REGION Network 16: TBD Stacking_New : Control Balize
   RUNG wire#powerrail
      Contact( "DB_MDM_SN".Energie )
      wire#w1
      Coil( #SN_bsr )
      Coil( "SN_Baliza dulap rosu" )
   END_RUNG
   RUNG wire#powerrail
      Contact( "DB_MDM_SN".No_Safe )
   END_RUNG wire#w1
   RUNG wire#powerrail
      Contact( "Gen".SN_AlarmAny )
   END_RUNG wire#w1
   RUNG wire#powerrail
      { S7_Templates := "SrcType := USInt" } EQ_Contact(in1 := "sn".f[5]."step", in2 := 2)
      wire#w2
      Contact( "DB2_WORK_BITS".Stacker_New_Handler.Input.Vertical_sus )
      Contact( "DB2_WORK_BITS".Stacker_New_Handler.Input.Furca_extins )
      Coil( #SN_bsy )
   END_RUNG
   RUNG wire#powerrail
      { S7_Templates := "SrcType := USInt" } EQ_Contact(in1 := "sn".f[5]."step", in2 := 4)
   END_RUNG wire#w2
   RUNG wire#powerrail
      I_Contact( "DB_MDM_SN".Energie )
      I_Contact( "DB_MDM_SN".No_Safe )
      I_Contact( "DB_MDM_SN".Cycle_Run )
      Coil( #SN_bsgc )
   END_RUNG
   RUNG wire#powerrail
      Contact( #SN_bsgc )
      Contact( "Clock_0.5Hz" )
      wire#w3
      Coil( "Sn_Baliza dulap verde" )
   END_RUNG
   RUNG wire#powerrail
      Contact( "DB_MDM_SN".Cycle_Run )
   END_RUNG wire#w3
   RUNG wire#w3
      Coil( #SN_bsg )
   END_RUNG
   RUNG wire#powerrail
      Contact( #SN_bsg )
      I_Contact( #SN_bsgc )
      Contact( #SN_bsy )
      Contact( "Clock_0.5Hz" )
      wire#w4
      Coil( "BS_G" )
   END_RUNG
   RUNG wire#powerrail
      Contact( #SN_bsg )
      I_Contact( #SN_bsy )
   END_RUNG wire#w4
   RUNG wire#powerrail
      Contact( #SN_bsg )
      Contact( #SN_bsy )
      wire#w5
      I_Contact( "Clock_0.5Hz" )
      Coil( "BS_Y" )
   END_RUNG
   RUNG wire#powerrail
      Contact( #SN_bsgc )
      Contact( #SN_bsy )
   END_RUNG wire#w5
   RUNG wire#powerrail
      Contact( #SN_bsr )
      Contact( #SN_bsy )
   END_RUNG wire#w5
   RUNG wire#powerrail
      Contact( #SN_bsr )
      wire#w6
      Contact( #SN_bsy )
      Contact( "Clock_0.5Hz" )
      wire#w7
      Coil( "BS_R" )
   END_RUNG
   RUNG wire#w6
      I_Contact( #SN_bsy )
   END_RUNG wire#w7
   // the same network as SCL:
   #SN_bsr := "DB_MDM_SN".Energie OR "DB_MDM_SN".No_Safe OR "Gen".SN_AlarmAny;
   "SN_Baliza dulap rosu" := #SN_bsr;
   #SN_bsy := (("sn".f[5]."step" = 2) OR ("sn".f[5]."step" = 4)) AND "DB2_WORK_BITS".Stacker_New_Handler.Input.Vertical_sus AND "DB2_WORK_BITS".Stacker_New_Handler.Input.Furca_extins;
   #SN_bsgc := NOT "DB_MDM_SN".Energie AND NOT "DB_MDM_SN".No_Safe AND NOT "DB_MDM_SN".Cycle_Run;
   "Sn_Baliza dulap verde" := (#SN_bsgc AND "Clock_0.5Hz") OR "DB_MDM_SN".Cycle_Run;
   #SN_bsg := "Sn_Baliza dulap verde";
   "BS_G" := (#SN_bsg AND NOT #SN_bsgc AND #SN_bsy AND "Clock_0.5Hz") OR (#SN_bsg AND NOT #SN_bsy);
   "BS_Y" := ((#SN_bsg AND #SN_bsy) OR (#SN_bsgc AND #SN_bsy) OR (#SN_bsr AND #SN_bsy)) AND NOT "Clock_0.5Hz";
   "BS_R" := #SN_bsr AND ((#SN_bsy AND "Clock_0.5Hz") OR NOT #SN_bsy);
END_REGION
END_FUNCTION

FUNCTION "FC20_HMI" : Void   // FC20, LAD
{ S7_Optimized_Access := 'TRUE' }
VERSION : 0.1
BEGIN

REGION Network 1
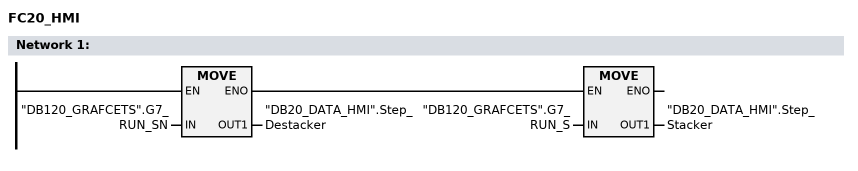
   RUNG wire#powerrail
      Move(in := "DB120_GRAFCETS".G7_RUN_SN, out1 => "DB20_DATA_HMI".Step_Destacker)
      Move(in := "DB120_GRAFCETS".G7_RUN_S, out1 => "DB20_DATA_HMI".Step_Stacker)
   END_RUNG
   // the same network as SCL:
   "DB20_DATA_HMI".Step_Destacker := "DB120_GRAFCETS".G7_RUN_SN;
   "DB20_DATA_HMI".Step_Stacker := "DB120_GRAFCETS".G7_RUN_S;
END_REGION
END_FUNCTION

FUNCTION "FC52_STACKING_New" : Void   // FC49, LAD
{ S7_Optimized_Access := 'TRUE' }
VERSION : 0.1
   VAR_TEMP
      Reset_S_Up : Bool;
      Reset_S_Fork : Bool;
      iB5_p : Bool;
      Reset_S : Bool;
      dumyb : Bool;
      dumyw : Int;
   END_VAR
   VAR_TEMP   // added for the SCL form of the ladder/FBD networks
      _w1 : Bool;
      _w2 : Bool;
      _w3 : Bool;
   END_VAR
BEGIN

REGION Network 1: mdm
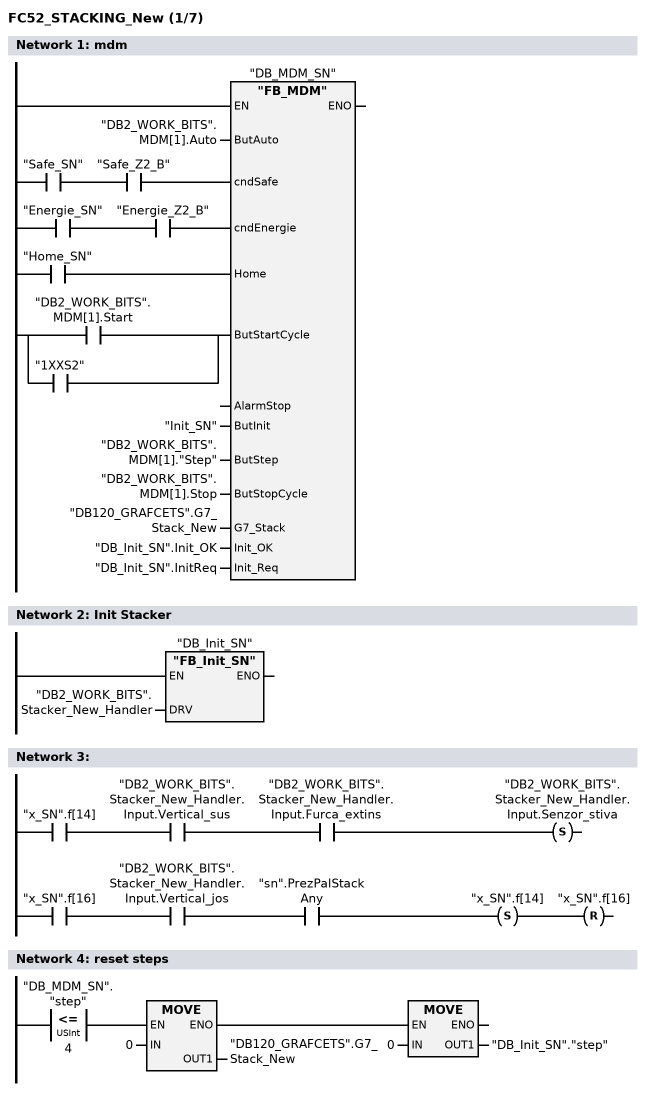
   RUNG wire#powerrail
      "DB_MDM_SN"(cndSafe := wire#w1, cndEnergie := wire#w2, Home := wire#w3, ButStartCycle := wire#w4, ButAuto := "DB2_WORK_BITS".MDM[1].Auto, AlarmStop :=, ButInit := "Init_SN", ButStep := "DB2_WORK_BITS".MDM[1]."Step", ButStopCycle := "DB2_WORK_BITS".MDM[1].Stop, G7_Stack := "DB120_GRAFCETS".G7_Stack_New, Init_OK := "DB_Init_SN".Init_OK, Init_Req := "DB_Init_SN".InitReq)
   END_RUNG
   RUNG wire#powerrail
      Contact( "Safe_SN" )
      Contact( "Safe_Z2_B" )
   END_RUNG wire#w1
   RUNG wire#powerrail
      Contact( "Energie_SN" )
      Contact( "Energie_Z2_B" )
   END_RUNG wire#w2
   RUNG wire#powerrail
      Contact( "Home_SN" )
   END_RUNG wire#w3
   RUNG wire#powerrail
      Contact( "DB2_WORK_BITS".MDM[1].Start )
   END_RUNG wire#w4
   RUNG wire#powerrail
      Contact( "1XXS2" )
   END_RUNG wire#w4
   // the same network as SCL:
   "DB_MDM_SN"(ButAuto := "DB2_WORK_BITS".MDM[1].Auto,   // "FB_MDM"
               cndSafe := "Safe_SN" AND "Safe_Z2_B",
               cndEnergie := "Energie_SN" AND "Energie_Z2_B",
               Home := "Home_SN",
               ButStartCycle := "DB2_WORK_BITS".MDM[1].Start OR "1XXS2",
               ButInit := "Init_SN",
               ButStep := "DB2_WORK_BITS".MDM[1]."Step",
               ButStopCycle := "DB2_WORK_BITS".MDM[1].Stop,
               G7_Stack := "DB120_GRAFCETS".G7_Stack_New,
               Init_OK := "DB_Init_SN".Init_OK,
               Init_Req := "DB_Init_SN".InitReq);
END_REGION

REGION Network 2: Init Stacker
   RUNG wire#powerrail
      "DB_Init_SN"(DRV := "DB2_WORK_BITS".Stacker_New_Handler)
   END_RUNG
   // the same network as SCL:
   "DB_Init_SN"(DRV := "DB2_WORK_BITS".Stacker_New_Handler);   // "FB_Init_SN"
END_REGION

REGION Network 3
   RUNG wire#powerrail
      Contact( "x_SN".f[14] )
      Contact( "DB2_WORK_BITS".Stacker_New_Handler.Input.Vertical_sus )
      Contact( "DB2_WORK_BITS".Stacker_New_Handler.Input.Furca_extins )
      S_Coil( "DB2_WORK_BITS".Stacker_New_Handler.Input.Senzor_stiva )
   END_RUNG
   RUNG wire#powerrail
      Contact( "x_SN".f[16] )
      Contact( "DB2_WORK_BITS".Stacker_New_Handler.Input.Vertical_jos )
      Contact( "sn".PrezPalStackAny )
      S_Coil( "x_SN".f[14] )
      R_Coil( "x_SN".f[16] )
   END_RUNG
   // the same network as SCL:
   IF "x_SN".f[14] AND "DB2_WORK_BITS".Stacker_New_Handler.Input.Vertical_sus AND "DB2_WORK_BITS".Stacker_New_Handler.Input.Furca_extins THEN
       "DB2_WORK_BITS".Stacker_New_Handler.Input.Senzor_stiva := TRUE;
   END_IF;
   #_w1 := "x_SN".f[16] AND "DB2_WORK_BITS".Stacker_New_Handler.Input.Vertical_jos AND "sn".PrezPalStackAny;
   IF #_w1 THEN
       "x_SN".f[14] := TRUE;
       "x_SN".f[16] := FALSE;
   END_IF;
END_REGION

REGION Network 4: reset steps
   RUNG wire#powerrail
      { S7_Templates := "SrcType := USInt" } LE_Contact(in1 := "DB_MDM_SN"."step", in2 := 4)
      Move(in := 0, out1 => "DB120_GRAFCETS".G7_Stack_New)
      Move(in := 0, out1 => "DB_Init_SN"."step")
   END_RUNG
   // the same network as SCL:
   IF "DB_MDM_SN"."step" <= 4 THEN
       "DB120_GRAFCETS".G7_Stack_New := 0;
       "DB_Init_SN"."step" := 0;
   END_IF;
END_REGION

REGION Network 5: start graf stack
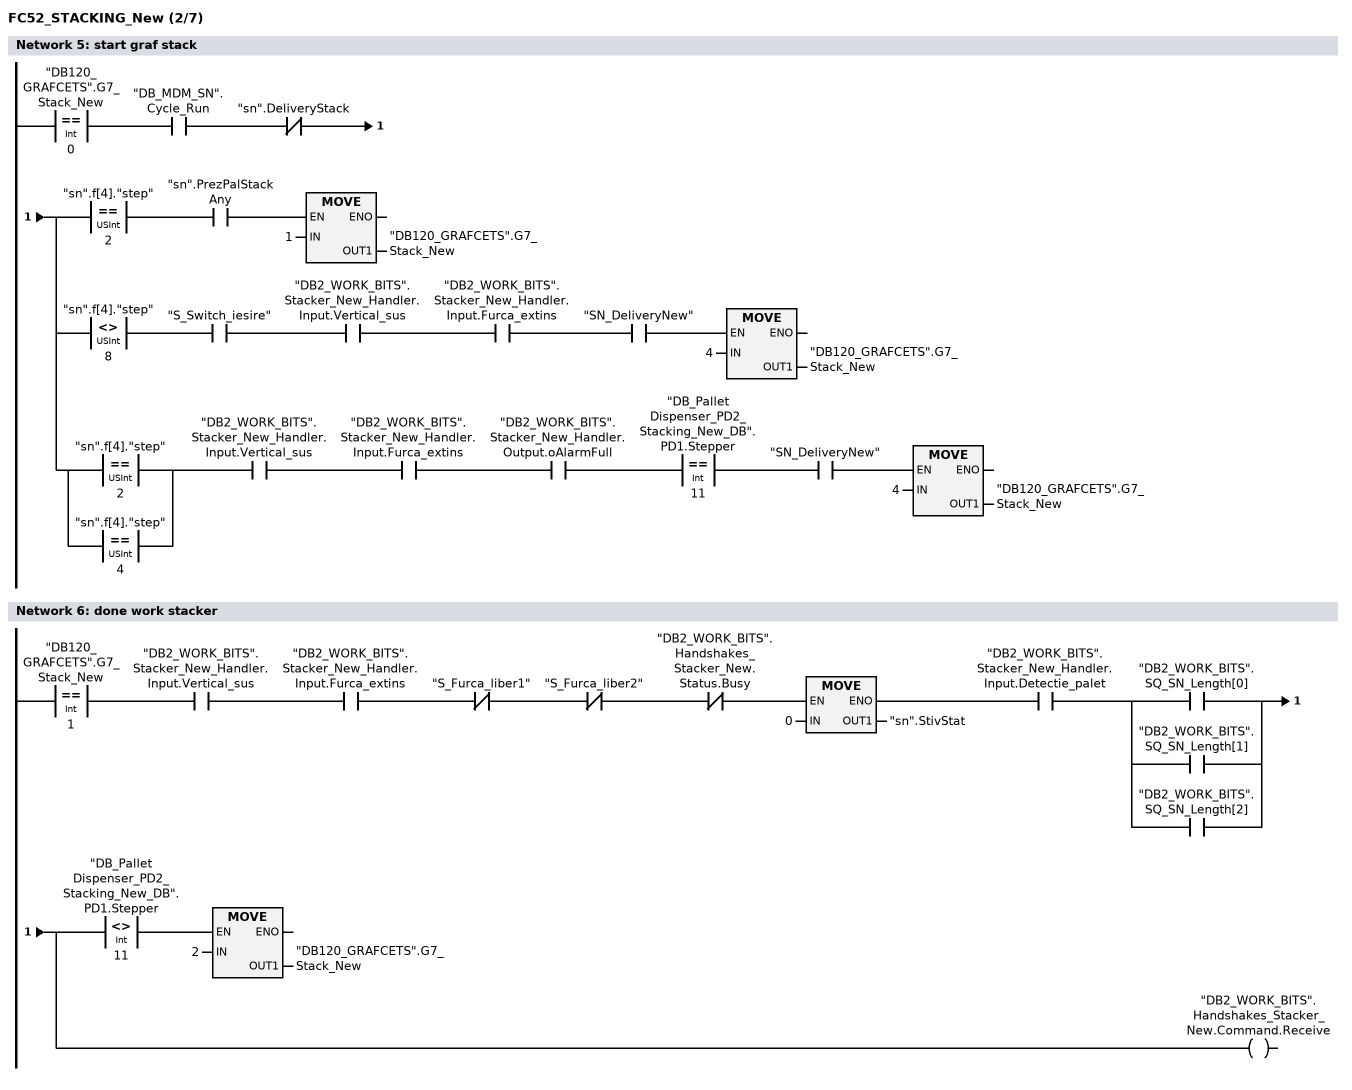
   RUNG wire#powerrail
      { S7_Templates := "SrcType := Int" } EQ_Contact(in1 := "DB120_GRAFCETS".G7_Stack_New, in2 := 0)
      Contact( "DB_MDM_SN".Cycle_Run )
      I_Contact( "sn".DeliveryStack )
      wire#w1
      { S7_Templates := "SrcType := USInt" } EQ_Contact(in1 := "sn".f[4]."step", in2 := 2)
      Contact( "sn".PrezPalStackAny )
      Move(in := 1, out1 => "DB120_GRAFCETS".G7_Stack_New)
   END_RUNG
   RUNG wire#w1
      { S7_Templates := "SrcType := USInt" } NE_Contact(in1 := "sn".f[4]."step", in2 := 8)
      Contact( "S_Switch_iesire" )
      Contact( "DB2_WORK_BITS".Stacker_New_Handler.Input.Vertical_sus )
      Contact( "DB2_WORK_BITS".Stacker_New_Handler.Input.Furca_extins )
      Contact( "SN_DeliveryNew" )
      Move(in := 4, out1 => "DB120_GRAFCETS".G7_Stack_New)
   END_RUNG
   RUNG wire#w1
      { S7_Templates := "SrcType := USInt" } EQ_Contact(in1 := "sn".f[4]."step", in2 := 2)
      wire#w2
      Contact( "DB2_WORK_BITS".Stacker_New_Handler.Input.Vertical_sus )
      Contact( "DB2_WORK_BITS".Stacker_New_Handler.Input.Furca_extins )
      Contact( "DB2_WORK_BITS".Stacker_New_Handler.Output.oAlarmFull )
      { S7_Templates := "SrcType := Int" } EQ_Contact(in1 := "DB_PalletDispenser_PD2_Stacking_New_DB".PD1.Stepper, in2 := 11)
      Contact( "SN_DeliveryNew" )
      Move(in := 4, out1 => "DB120_GRAFCETS".G7_Stack_New)
   END_RUNG
   RUNG wire#w1
      { S7_Templates := "SrcType := USInt" } EQ_Contact(in1 := "sn".f[4]."step", in2 := 4)
   END_RUNG wire#w2
   // the same network as SCL:
   #_w1 := ("DB120_GRAFCETS".G7_Stack_New = 0) AND "DB_MDM_SN".Cycle_Run AND NOT "sn".DeliveryStack;
   IF #_w1 AND ("sn".f[4]."step" = 2) AND "sn".PrezPalStackAny THEN
       "DB120_GRAFCETS".G7_Stack_New := 1;
   END_IF;
   IF #_w1 AND ("sn".f[4]."step" <> 8) AND "S_Switch_iesire" AND "DB2_WORK_BITS".Stacker_New_Handler.Input.Vertical_sus AND "DB2_WORK_BITS".Stacker_New_Handler.Input.Furca_extins AND "SN_DeliveryNew" THEN
       "DB120_GRAFCETS".G7_Stack_New := 4;
   END_IF;
   IF #_w1 AND (("sn".f[4]."step" = 2) OR ("sn".f[4]."step" = 4)) AND "DB2_WORK_BITS".Stacker_New_Handler.Input.Vertical_sus AND "DB2_WORK_BITS".Stacker_New_Handler.Input.Furca_extins AND "DB2_WORK_BITS".Stacker_New_Handler.Output.oAlarmFull AND ("DB_PalletDispenser_PD2_Stacking_New_DB".PD1.Stepper = 11) AND "SN_DeliveryNew" THEN
       "DB120_GRAFCETS".G7_Stack_New := 4;
   END_IF;
END_REGION

REGION Network 6: done work stacker
   RUNG wire#powerrail
      { S7_Templates := "SrcType := Int" } EQ_Contact(in1 := "DB120_GRAFCETS".G7_Stack_New, in2 := 1)
      Contact( "DB2_WORK_BITS".Stacker_New_Handler.Input.Vertical_sus )
      Contact( "DB2_WORK_BITS".Stacker_New_Handler.Input.Furca_extins )
      I_Contact( "S_Furca_liber1" )
      I_Contact( "S_Furca_liber2" )
      I_Contact( "DB2_WORK_BITS".Handshakes_Stacker_New.Status.Busy )
      Move(in := 0, out1 => "sn".StivStat)
      Contact( "DB2_WORK_BITS".Stacker_New_Handler.Input.Detectie_palet )
      wire#w1
      Contact( "DB2_WORK_BITS".SQ_SN_Length[0] )
      wire#w2
      { S7_Templates := "SrcType := Int" } NE_Contact(in1 := "DB_PalletDispenser_PD2_Stacking_New_DB".PD1.Stepper, in2 := 11)
      Move(in := 2, out1 => "DB120_GRAFCETS".G7_Stack_New)
   END_RUNG
   RUNG wire#w1
      Contact( "DB2_WORK_BITS".SQ_SN_Length[1] )
   END_RUNG wire#w2
   RUNG wire#w1
      Contact( "DB2_WORK_BITS".SQ_SN_Length[2] )
   END_RUNG wire#w2
   RUNG wire#w2
      Coil( "DB2_WORK_BITS".Handshakes_Stacker_New.Command.Receive )
   END_RUNG
   // the same network as SCL:
   #_w1 := ("DB120_GRAFCETS".G7_Stack_New = 1) AND "DB2_WORK_BITS".Stacker_New_Handler.Input.Vertical_sus AND "DB2_WORK_BITS".Stacker_New_Handler.Input.Furca_extins AND NOT "S_Furca_liber1" AND NOT "S_Furca_liber2" AND NOT "DB2_WORK_BITS".Handshakes_Stacker_New.Status.Busy;
   IF #_w1 THEN "sn".StivStat := 0; END_IF;
   #_w2 := #_w1 AND "DB2_WORK_BITS".Stacker_New_Handler.Input.Detectie_palet AND ("DB2_WORK_BITS".SQ_SN_Length[0] OR "DB2_WORK_BITS".SQ_SN_Length[1] OR "DB2_WORK_BITS".SQ_SN_Length[2]);
   IF #_w2 AND ("DB_PalletDispenser_PD2_Stacking_New_DB".PD1.Stepper <> 11) THEN
       "DB120_GRAFCETS".G7_Stack_New := 2;
   END_IF;
   "DB2_WORK_BITS".Handshakes_Stacker_New.Command.Receive := #_w2;
END_REGION

REGION Network 7: decision continue/release stack
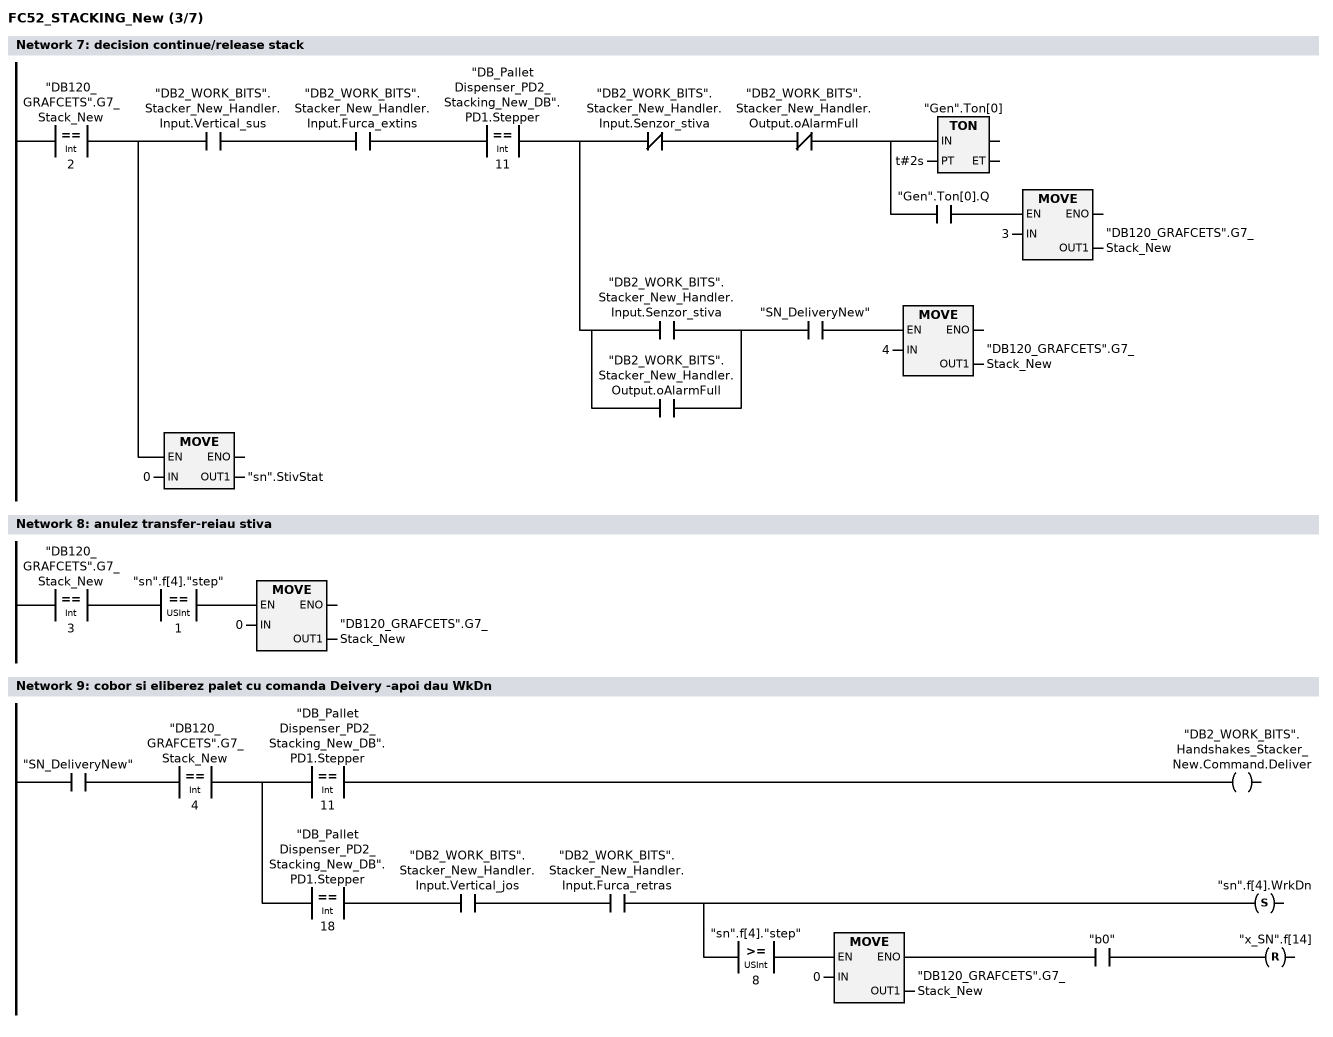
   #_w1 := "DB120_GRAFCETS".G7_Stack_New = 2;
   #_w2 := #_w1 AND "DB2_WORK_BITS".Stacker_New_Handler.Input.Vertical_sus AND "DB2_WORK_BITS".Stacker_New_Handler.Input.Furca_extins AND ("DB_PalletDispenser_PD2_Stacking_New_DB".PD1.Stepper = 11);
   #_w3 := #_w2 AND NOT "DB2_WORK_BITS".Stacker_New_Handler.Input.Senzor_stiva AND NOT "DB2_WORK_BITS".Stacker_New_Handler.Output.oAlarmFull;
   "Gen".Ton[0].TON(IN := #_w3, PT := t#2s);
   IF #_w3 AND "Gen".Ton[0].Q THEN "DB120_GRAFCETS".G7_Stack_New := 3; END_IF;
   IF #_w2 AND ("DB2_WORK_BITS".Stacker_New_Handler.Input.Senzor_stiva OR "DB2_WORK_BITS".Stacker_New_Handler.Output.oAlarmFull) AND "SN_DeliveryNew" THEN
       "DB120_GRAFCETS".G7_Stack_New := 4;
   END_IF;
   IF #_w1 THEN "sn".StivStat := 0; END_IF;
END_REGION

REGION Network 8: anulez transfer-reiau stiva
   RUNG wire#powerrail
      { S7_Templates := "SrcType := Int" } EQ_Contact(in1 := "DB120_GRAFCETS".G7_Stack_New, in2 := 3)
      { S7_Templates := "SrcType := USInt" } EQ_Contact(in1 := "sn".f[4]."step", in2 := 1)
      Move(in := 0, out1 => "DB120_GRAFCETS".G7_Stack_New)
   END_RUNG
   // the same network as SCL:
   IF ("DB120_GRAFCETS".G7_Stack_New = 3) AND ("sn".f[4]."step" = 1) THEN
       "DB120_GRAFCETS".G7_Stack_New := 0;
   END_IF;
END_REGION

REGION Network 9: cobor si eliberez palet cu comanda Deivery -apoi dau WkDn
   RUNG wire#powerrail
      Contact( "SN_DeliveryNew" )
      { S7_Templates := "SrcType := Int" } EQ_Contact(in1 := "DB120_GRAFCETS".G7_Stack_New, in2 := 4)
      wire#w1
      { S7_Templates := "SrcType := Int" } EQ_Contact(in1 := "DB_PalletDispenser_PD2_Stacking_New_DB".PD1.Stepper, in2 := 11)
      Coil( "DB2_WORK_BITS".Handshakes_Stacker_New.Command.Deliver )
   END_RUNG
   RUNG wire#w1
      { S7_Templates := "SrcType := Int" } EQ_Contact(in1 := "DB_PalletDispenser_PD2_Stacking_New_DB".PD1.Stepper, in2 := 18)
      Contact( "DB2_WORK_BITS".Stacker_New_Handler.Input.Vertical_jos )
      Contact( "DB2_WORK_BITS".Stacker_New_Handler.Input.Furca_retras )
      wire#w2
      S_Coil( "sn".f[4].WrkDn )
   END_RUNG
   RUNG wire#w2
      { S7_Templates := "SrcType := USInt" } GE_Contact(in1 := "sn".f[4]."step", in2 := 8)
      Move(in := 0, out1 => "DB120_GRAFCETS".G7_Stack_New)
      Contact( "b0" )
      R_Coil( "x_SN".f[14] )
   END_RUNG
   // the same network as SCL:
   #_w1 := "SN_DeliveryNew" AND ("DB120_GRAFCETS".G7_Stack_New = 4);
   "DB2_WORK_BITS".Handshakes_Stacker_New.Command.Deliver := #_w1 AND ("DB_PalletDispenser_PD2_Stacking_New_DB".PD1.Stepper = 11);
   #_w2 := #_w1 AND ("DB_PalletDispenser_PD2_Stacking_New_DB".PD1.Stepper = 18) AND "DB2_WORK_BITS".Stacker_New_Handler.Input.Vertical_jos AND "DB2_WORK_BITS".Stacker_New_Handler.Input.Furca_retras;
   IF #_w2 THEN "sn".f[4].WrkDn := TRUE; END_IF;
   #_w3 := #_w2 AND ("sn".f[4]."step" >= 8);
   IF #_w3 THEN "DB120_GRAFCETS".G7_Stack_New := 0; END_IF;
   IF #_w3 AND "b0" THEN "x_SN".f[14] := FALSE; END_IF;
END_REGION

REGION Network 10: delivery
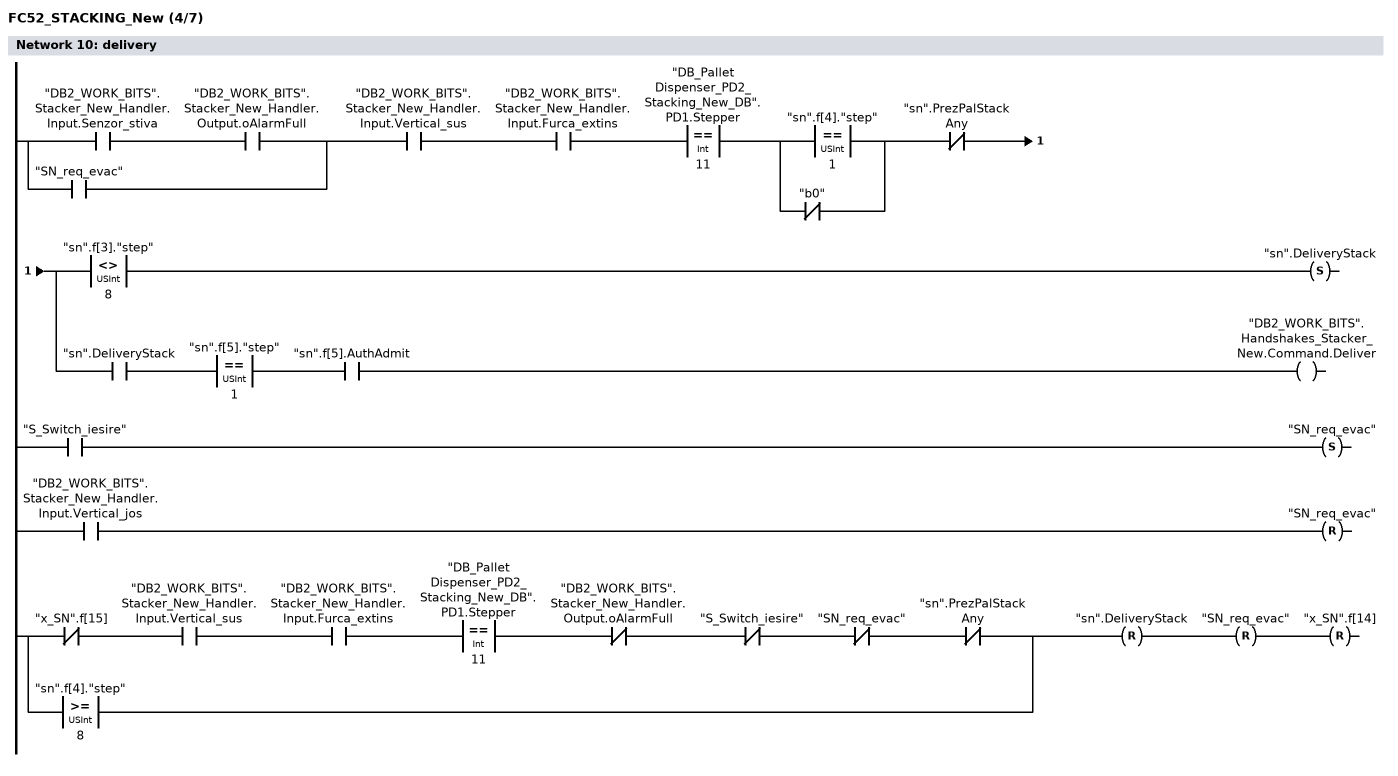
   RUNG wire#powerrail
      Contact( "DB2_WORK_BITS".Stacker_New_Handler.Input.Senzor_stiva )
      Contact( "DB2_WORK_BITS".Stacker_New_Handler.Output.oAlarmFull )
      wire#w1
      Contact( "DB2_WORK_BITS".Stacker_New_Handler.Input.Vertical_sus )
      Contact( "DB2_WORK_BITS".Stacker_New_Handler.Input.Furca_extins )
      { S7_Templates := "SrcType := Int" } EQ_Contact(in1 := "DB_PalletDispenser_PD2_Stacking_New_DB".PD1.Stepper, in2 := 11)
      wire#w2
      { S7_Templates := "SrcType := USInt" } EQ_Contact(in1 := "sn".f[4]."step", in2 := 1)
      wire#w3
      I_Contact( "sn".PrezPalStackAny )
      wire#w4
      { S7_Templates := "SrcType := USInt" } NE_Contact(in1 := "sn".f[3]."step", in2 := 8)
      S_Coil( "sn".DeliveryStack )
   END_RUNG
   RUNG wire#powerrail
      Contact( "SN_req_evac" )
   END_RUNG wire#w1
   RUNG wire#w2
      I_Contact( "b0" )
   END_RUNG wire#w3
   RUNG wire#w4
      Contact( "sn".DeliveryStack )
      { S7_Templates := "SrcType := USInt" } EQ_Contact(in1 := "sn".f[5]."step", in2 := 1)
      Contact( "sn".f[5].AuthAdmit )
      Coil( "DB2_WORK_BITS".Handshakes_Stacker_New.Command.Deliver )
   END_RUNG
   RUNG wire#powerrail
      Contact( "S_Switch_iesire" )
      S_Coil( "SN_req_evac" )
   END_RUNG
   RUNG wire#powerrail
      Contact( "DB2_WORK_BITS".Stacker_New_Handler.Input.Vertical_jos )
      R_Coil( "SN_req_evac" )
   END_RUNG
   RUNG wire#powerrail
      I_Contact( "x_SN".f[15] )
      Contact( "DB2_WORK_BITS".Stacker_New_Handler.Input.Vertical_sus )
      Contact( "DB2_WORK_BITS".Stacker_New_Handler.Input.Furca_extins )
      { S7_Templates := "SrcType := Int" } EQ_Contact(in1 := "DB_PalletDispenser_PD2_Stacking_New_DB".PD1.Stepper, in2 := 11)
      I_Contact( "DB2_WORK_BITS".Stacker_New_Handler.Output.oAlarmFull )
      I_Contact( "S_Switch_iesire" )
      I_Contact( "SN_req_evac" )
      I_Contact( "sn".PrezPalStackAny )
      wire#w5
      R_Coil( "sn".DeliveryStack )
      R_Coil( "SN_req_evac" )
      R_Coil( "x_SN".f[14] )
   END_RUNG
   RUNG wire#powerrail
      { S7_Templates := "SrcType := USInt" } GE_Contact(in1 := "sn".f[4]."step", in2 := 8)
   END_RUNG wire#w5
   // the same network as SCL:
   #_w1 := (("DB2_WORK_BITS".Stacker_New_Handler.Input.Senzor_stiva AND "DB2_WORK_BITS".Stacker_New_Handler.Output.oAlarmFull) OR "SN_req_evac") AND "DB2_WORK_BITS".Stacker_New_Handler.Input.Vertical_sus AND "DB2_WORK_BITS".Stacker_New_Handler.Input.Furca_extins AND ("DB_PalletDispenser_PD2_Stacking_New_DB".PD1.Stepper = 11) AND (("sn".f[4]."step" = 1) OR NOT "b0") AND NOT "sn".PrezPalStackAny;
   IF #_w1 AND ("sn".f[3]."step" <> 8) THEN "sn".DeliveryStack := TRUE; END_IF;
   "DB2_WORK_BITS".Handshakes_Stacker_New.Command.Deliver := #_w1 AND "sn".DeliveryStack AND ("sn".f[5]."step" = 1) AND "sn".f[5].AuthAdmit;
   IF "S_Switch_iesire" THEN "SN_req_evac" := TRUE; END_IF;
   IF "DB2_WORK_BITS".Stacker_New_Handler.Input.Vertical_jos THEN "SN_req_evac" := FALSE; END_IF;
   IF (NOT "x_SN".f[15] AND "DB2_WORK_BITS".Stacker_New_Handler.Input.Vertical_sus AND "DB2_WORK_BITS".Stacker_New_Handler.Input.Furca_extins AND ("DB_PalletDispenser_PD2_Stacking_New_DB".PD1.Stepper = 11) AND NOT "DB2_WORK_BITS".Stacker_New_Handler.Output.oAlarmFull AND NOT "S_Switch_iesire" AND NOT "SN_req_evac" AND NOT "sn".PrezPalStackAny) OR ("sn".f[4]."step" >= 8) THEN
       "sn".DeliveryStack := FALSE;
   END_IF;
   #_w2 := (NOT "x_SN".f[15] AND "DB2_WORK_BITS".Stacker_New_Handler.Input.Vertical_sus AND "DB2_WORK_BITS".Stacker_New_Handler.Input.Furca_extins AND ("DB_PalletDispenser_PD2_Stacking_New_DB".PD1.Stepper = 11) AND NOT "DB2_WORK_BITS".Stacker_New_Handler.Output.oAlarmFull AND NOT "S_Switch_iesire" AND NOT "SN_req_evac" AND NOT "sn".PrezPalStackAny) OR ("sn".f[4]."step" >= 8);
   IF #_w2 THEN
       "SN_req_evac" := FALSE;
       "x_SN".f[14] := FALSE;
   END_IF;
END_REGION

REGION Network 11: call FB stack
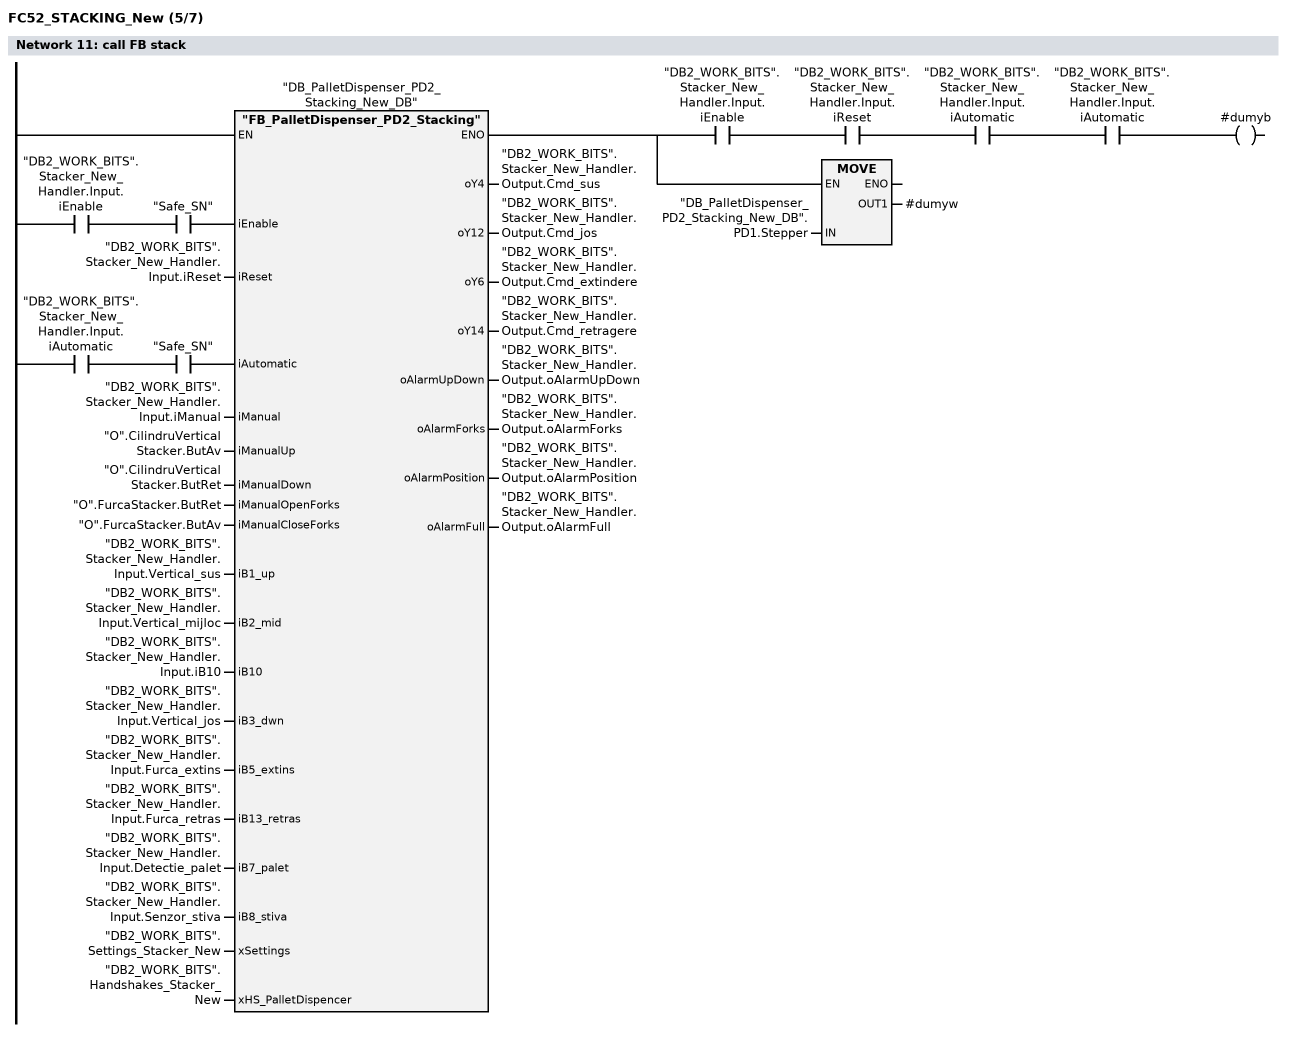
   RUNG wire#powerrail
      "DB_PalletDispenser_PD2_Stacking_New_DB"(iEnable := wire#w1, iAutomatic := wire#w2, iReset := "DB2_WORK_BITS".Stacker_New_Handler.Input.iReset, iManual := "DB2_WORK_BITS".Stacker_New_Handler.Input.iManual, iManualUp := "O".CilindruVerticalStacker.ButAv, iManualDown := "O".CilindruVerticalStacker.ButRet, iManualOpenForks := "O".FurcaStacker.ButRet, iManualCloseForks := "O".FurcaStacker.ButAv, iB1_up := "DB2_WORK_BITS".Stacker_New_Handler.Input.Vertical_sus, iB2_mid := "DB2_WORK_BITS".Stacker_New_Handler.Input.Vertical_mijloc, iB10 := "DB2_WORK_BITS".Stacker_New_Handler.Input.iB10, iB3_dwn := "DB2_WORK_BITS".Stacker_New_Handler.Input.Vertical_jos, iB5_extins := "DB2_WORK_BITS".Stacker_New_Handler.Input.Furca_extins, iB13_retras := "DB2_WORK_BITS".Stacker_New_Handler.Input.Furca_retras, iB7_palet := "DB2_WORK_BITS".Stacker_New_Handler.Input.Detectie_palet, iB8_stiva := "DB2_WORK_BITS".Stacker_New_Handler.Input.Senzor_stiva, xSettings := "DB2_WORK_BITS".Settings_Stacker_New, xHS_PalletDispencer := "DB2_WORK_BITS".Handshakes_Stacker_New, oY4 => "DB2_WORK_BITS".Stacker_New_Handler.Output.Cmd_sus, oY12 => "DB2_WORK_BITS".Stacker_New_Handler.Output.Cmd_jos, oY6 => "DB2_WORK_BITS".Stacker_New_Handler.Output.Cmd_extindere, oY14 => "DB2_WORK_BITS".Stacker_New_Handler.Output.Cmd_retragere, oAlarmUpDown => "DB2_WORK_BITS".Stacker_New_Handler.Output.oAlarmUpDown, oAlarmForks => "DB2_WORK_BITS".Stacker_New_Handler.Output.oAlarmForks, oAlarmPosition => "DB2_WORK_BITS".Stacker_New_Handler.Output.oAlarmPosition, oAlarmFull => "DB2_WORK_BITS".Stacker_New_Handler.Output.oAlarmFull)
      wire#w3
      Contact( "DB2_WORK_BITS".Stacker_New_Handler.Input.iEnable )
      Contact( "DB2_WORK_BITS".Stacker_New_Handler.Input.iReset )
      Contact( "DB2_WORK_BITS".Stacker_New_Handler.Input.iAutomatic )
      Contact( "DB2_WORK_BITS".Stacker_New_Handler.Input.iAutomatic )
      Coil( #dumyb )
   END_RUNG
   RUNG wire#powerrail
      Contact( "DB2_WORK_BITS".Stacker_New_Handler.Input.iEnable )
      Contact( "Safe_SN" )
   END_RUNG wire#w1
   RUNG wire#powerrail
      Contact( "DB2_WORK_BITS".Stacker_New_Handler.Input.iAutomatic )
      Contact( "Safe_SN" )
   END_RUNG wire#w2
   RUNG wire#w3
      Move(in := "DB_PalletDispenser_PD2_Stacking_New_DB".PD1.Stepper, out1 => #dumyw)
   END_RUNG
   // the same network as SCL:
   "DB_PalletDispenser_PD2_Stacking_New_DB"(iEnable := "DB2_WORK_BITS".Stacker_New_Handler.Input.iEnable AND "Safe_SN",   // "FB_PalletDispenser_PD2_Stacking"
                           iReset := "DB2_WORK_BITS".Stacker_New_Handler.Input.iReset,
                           iAutomatic := "DB2_WORK_BITS".Stacker_New_Handler.Input.iAutomatic AND "Safe_SN",
                           iManual := "DB2_WORK_BITS".Stacker_New_Handler.Input.iManual,
                           iManualUp := "O".CilindruVerticalStacker.ButAv,
                           iManualDown := "O".CilindruVerticalStacker.ButRet,
                           iManualOpenForks := "O".FurcaStacker.ButRet,
                           iManualCloseForks := "O".FurcaStacker.ButAv,
                           iB1_up := "DB2_WORK_BITS".Stacker_New_Handler.Input.Vertical_sus,
                           iB2_mid := "DB2_WORK_BITS".Stacker_New_Handler.Input.Vertical_mijloc,
                           iB10 := "DB2_WORK_BITS".Stacker_New_Handler.Input.iB10,
                           iB3_dwn := "DB2_WORK_BITS".Stacker_New_Handler.Input.Vertical_jos,
                           iB5_extins := "DB2_WORK_BITS".Stacker_New_Handler.Input.Furca_extins,
                           iB13_retras := "DB2_WORK_BITS".Stacker_New_Handler.Input.Furca_retras,
                           iB7_palet := "DB2_WORK_BITS".Stacker_New_Handler.Input.Detectie_palet,
                           iB8_stiva := "DB2_WORK_BITS".Stacker_New_Handler.Input.Senzor_stiva,
                           xSettings := "DB2_WORK_BITS".Settings_Stacker_New,
                           xHS_PalletDispencer := "DB2_WORK_BITS".Handshakes_Stacker_New,
                           oY4 => "DB2_WORK_BITS".Stacker_New_Handler.Output.Cmd_sus,
                           oY12 => "DB2_WORK_BITS".Stacker_New_Handler.Output.Cmd_jos,
                           oY6 => "DB2_WORK_BITS".Stacker_New_Handler.Output.Cmd_extindere,
                           oY14 => "DB2_WORK_BITS".Stacker_New_Handler.Output.Cmd_retragere,
                           oAlarmUpDown => "DB2_WORK_BITS".Stacker_New_Handler.Output.oAlarmUpDown,
                           oAlarmForks => "DB2_WORK_BITS".Stacker_New_Handler.Output.oAlarmForks,
                           oAlarmPosition => "DB2_WORK_BITS".Stacker_New_Handler.Output.oAlarmPosition,
                           oAlarmFull => "DB2_WORK_BITS".Stacker_New_Handler.Output.oAlarmFull,
                           ENO => #_w1);
   #dumyb := #_w1 AND "DB2_WORK_BITS".Stacker_New_Handler.Input.iEnable AND "DB2_WORK_BITS".Stacker_New_Handler.Input.iReset AND "DB2_WORK_BITS".Stacker_New_Handler.Input.iAutomatic AND "DB2_WORK_BITS".Stacker_New_Handler.Input.iAutomatic;
   IF #_w1 THEN #dumyw := "DB_PalletDispenser_PD2_Stacking_New_DB".PD1.Stepper; END_IF;
END_REGION

REGION Network 12: iEnable
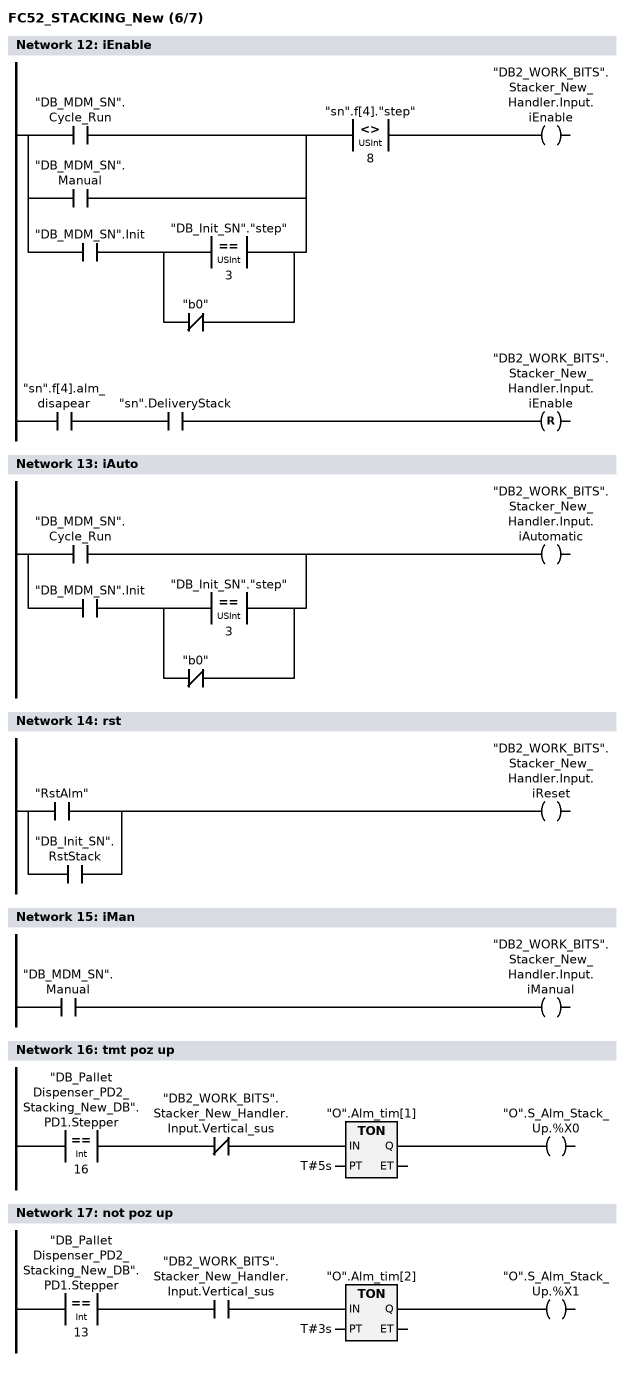
   RUNG wire#powerrail
      Contact( "DB_MDM_SN".Cycle_Run )
      wire#w1
      { S7_Templates := "SrcType := USInt" } NE_Contact(in1 := "sn".f[4]."step", in2 := 8)
      Coil( "DB2_WORK_BITS".Stacker_New_Handler.Input.iEnable )
   END_RUNG
   RUNG wire#powerrail
      Contact( "DB_MDM_SN".Manual )
   END_RUNG wire#w1
   RUNG wire#powerrail
      Contact( "DB_MDM_SN".Init )
      wire#w2
      { S7_Templates := "SrcType := USInt" } EQ_Contact(in1 := "DB_Init_SN"."step", in2 := 3)
   END_RUNG wire#w1
   RUNG wire#w2
      I_Contact( "b0" )
   END_RUNG wire#w1
   RUNG wire#powerrail
      Contact( "sn".f[4].alm_disapear )
      Contact( "sn".DeliveryStack )
      R_Coil( "DB2_WORK_BITS".Stacker_New_Handler.Input.iEnable )
   END_RUNG
   // the same network as SCL:
   "DB2_WORK_BITS".Stacker_New_Handler.Input.iEnable := ("DB_MDM_SN".Cycle_Run OR "DB_MDM_SN".Manual OR ("DB_MDM_SN".Init AND (("DB_Init_SN"."step" = 3) OR NOT "b0"))) AND ("sn".f[4]."step" <> 8);
   IF "sn".f[4].alm_disapear AND "sn".DeliveryStack THEN
       "DB2_WORK_BITS".Stacker_New_Handler.Input.iEnable := FALSE;
   END_IF;
END_REGION

REGION Network 13: iAuto
   RUNG wire#powerrail
      Contact( "DB_MDM_SN".Cycle_Run )
      wire#w1
      Coil( "DB2_WORK_BITS".Stacker_New_Handler.Input.iAutomatic )
   END_RUNG
   RUNG wire#powerrail
      Contact( "DB_MDM_SN".Init )
      wire#w2
      { S7_Templates := "SrcType := USInt" } EQ_Contact(in1 := "DB_Init_SN"."step", in2 := 3)
   END_RUNG wire#w1
   RUNG wire#w2
      I_Contact( "b0" )
   END_RUNG wire#w1
   // the same network as SCL:
   "DB2_WORK_BITS".Stacker_New_Handler.Input.iAutomatic := "DB_MDM_SN".Cycle_Run OR ("DB_MDM_SN".Init AND (("DB_Init_SN"."step" = 3) OR NOT "b0"));
END_REGION

REGION Network 14: rst
   RUNG wire#powerrail
      Contact( "RstAlm" )
      wire#w1
      Coil( "DB2_WORK_BITS".Stacker_New_Handler.Input.iReset )
   END_RUNG
   RUNG wire#powerrail
      Contact( "DB_Init_SN".RstStack )
   END_RUNG wire#w1
   // the same network as SCL:
   "DB2_WORK_BITS".Stacker_New_Handler.Input.iReset := "RstAlm" OR "DB_Init_SN".RstStack;
END_REGION

REGION Network 15: iMan
   RUNG wire#powerrail
      Contact( "DB_MDM_SN".Manual )
      Coil( "DB2_WORK_BITS".Stacker_New_Handler.Input.iManual )
   END_RUNG
   // the same network as SCL:
   "DB2_WORK_BITS".Stacker_New_Handler.Input.iManual := "DB_MDM_SN".Manual;
END_REGION

REGION Network 16: tmt poz up
   "O".Alm_tim[1].TON(IN := ("DB_PalletDispenser_PD2_Stacking_New_DB".PD1.Stepper = 16) AND NOT "DB2_WORK_BITS".Stacker_New_Handler.Input.Vertical_sus,
                      PT := T#5s);
   "O".S_Alm_Stack_Up.%X0 := "O".Alm_tim[1].Q;
END_REGION

REGION Network 17: not poz up
   "O".Alm_tim[2].TON(IN := ("DB_PalletDispenser_PD2_Stacking_New_DB".PD1.Stepper = 13) AND "DB2_WORK_BITS".Stacker_New_Handler.Input.Vertical_sus,
                      PT := T#3s);
   "O".S_Alm_Stack_Up.%X1 := "O".Alm_tim[2].Q;
END_REGION

REGION Network 18: lose poz up
